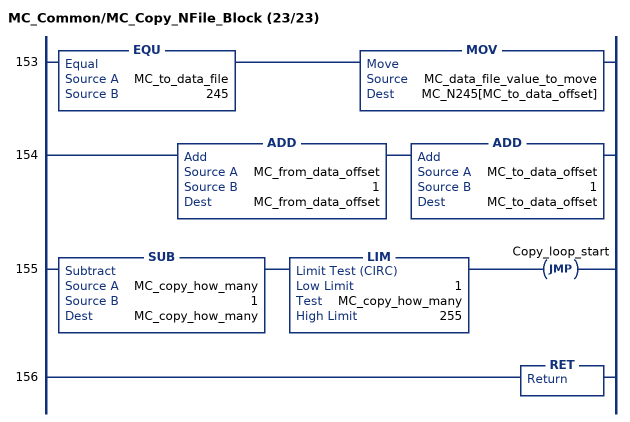
   153: EQU(MC_to_data_file,245)MOV(MC_data_file_value_to_move,MC_N245[MC_to_data_offset]);
   154: ADD(MC_from_data_offset,1,MC_from_data_offset)ADD(MC_to_data_offset,1,MC_to_data_offset);
   155: SUB(MC_copy_how_many,1,MC_copy_how_many)LIM(1,MC_copy_how_many,255)JMP(Copy_loop_start);
   156: RET();
END_ROUTINE

ROUTINE MC_DEBOUNCE_3   (* ladder *)
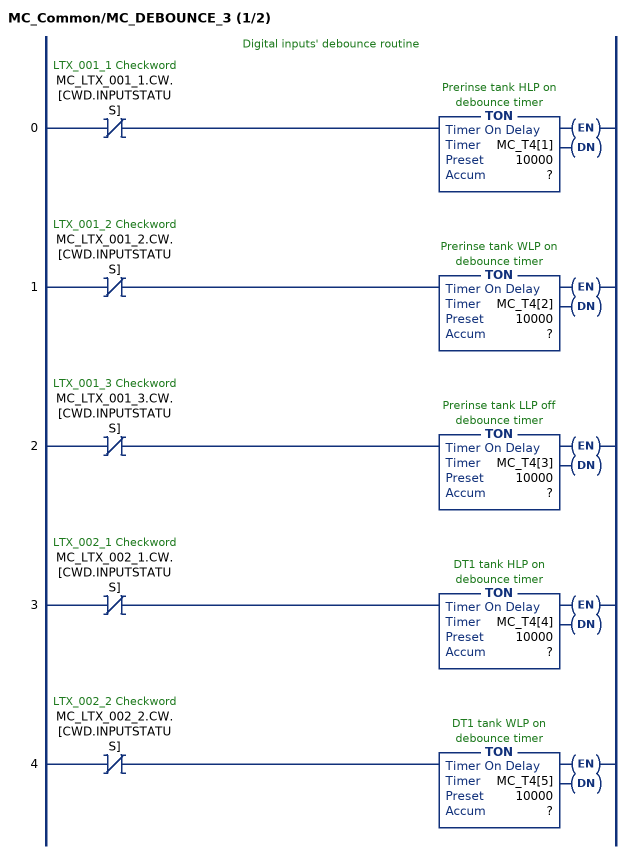
   // Digital inputs' debounce routine
   0: XIO(MC_LTX_001_1.CW.[CWD.INPUTSTATUS])TON(MC_T4[1],?,?);
   1: XIO(MC_LTX_001_2.CW.[CWD.INPUTSTATUS])TON(MC_T4[2],?,?);
   2: XIO(MC_LTX_001_3.CW.[CWD.INPUTSTATUS])TON(MC_T4[3],?,?);
   3: XIO(MC_LTX_002_1.CW.[CWD.INPUTSTATUS])TON(MC_T4[4],?,?);
   4: XIO(MC_LTX_002_2.CW.[CWD.INPUTSTATUS])TON(MC_T4[5],?,?);
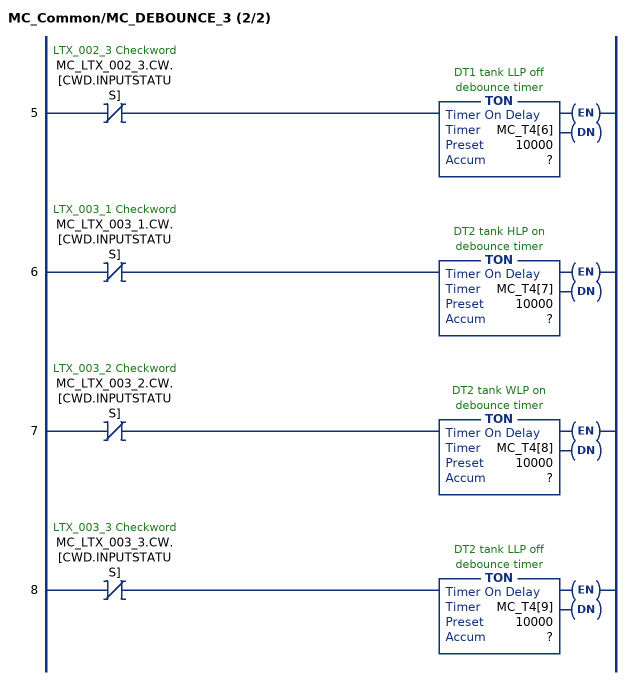
   5: XIO(MC_LTX_002_3.CW.[CWD.INPUTSTATUS])TON(MC_T4[6],?,?);
   6: XIO(MC_LTX_003_1.CW.[CWD.INPUTSTATUS])TON(MC_T4[7],?,?);
   7: XIO(MC_LTX_003_2.CW.[CWD.INPUTSTATUS])TON(MC_T4[8],?,?);
   8: XIO(MC_LTX_003_3.CW.[CWD.INPUTSTATUS])TON(MC_T4[9],?,?);
END_ROUTINE

ROUTINE MC_Digital_Inputs   (* ladder *)
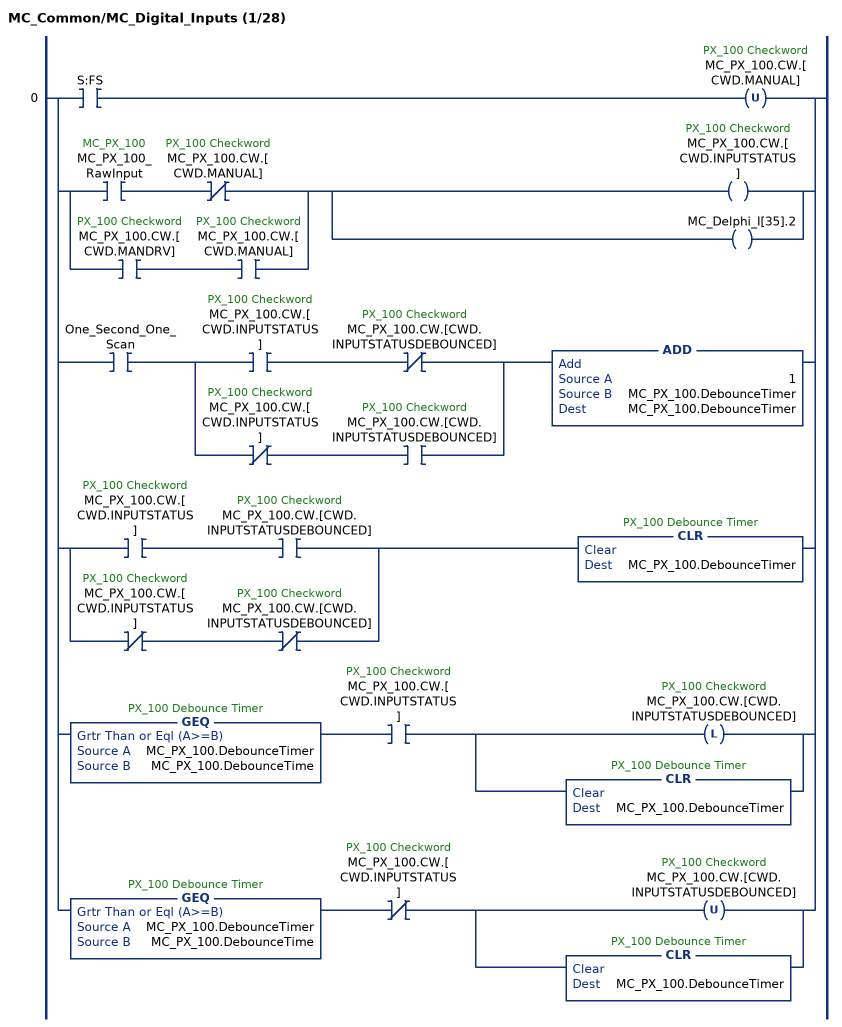
   0: [XIC(S:FS) OTU(MC_PX_100.CW.[CWD.MANUAL]) ,[XIC(MC_PX_100_RawInput) XIO(MC_PX_100.CW.[CWD.MANUAL]) ,XIC(MC_PX_100.CW.[CWD.MANDRV]) XIC(MC_PX_100.CW.[CWD.MANUAL]) ] [OTE(MC_PX_100.CW.[CWD.INPUTSTATUS]) ,OTE(MC_Delphi_I[35].2) ] ,XIC(One_Second_One_Scan) [XIC(MC_PX_100.CW.[CWD.INPUTSTATUS]) XIO(MC_PX_100.CW.[CWD.INPUTSTATUSDEBOUNCED]) ,XIO(MC_PX_100.CW.[CWD.INPUTSTATUS]) XIC(MC_PX_100.CW.[CWD.INPUTSTATUSDEBOUNCED]) ] ADD(1,MC_PX_100.DebounceTimer,MC_PX_100.DebounceTimer) ,[XIC(MC_PX_100.CW.[CWD.INPUTSTATUS]) XIC(MC_PX_100.CW.[CWD.INPUTSTATUSDEBOUNCED]) ,XIO(MC_PX_100.CW.[CWD.INPUTSTATUS]) XIO(MC_PX_100.CW.[CWD.INPUTSTATUSDEBOUNCED]) ] CLR(MC_PX_100.DebounceTimer) ,GEQ(MC_PX_100.DebounceTimer,MC_PX_100.DebounceTime) XIC(MC_PX_100.CW.[CWD.INPUTSTATUS]) [OTL(MC_PX_100.CW.[CWD.INPUTSTATUSDEBOUNCED]) ,CLR(MC_PX_100.DebounceTimer) ] ,GEQ(MC_PX_100.DebounceTimer,MC_PX_100.DebounceTime) XIO(MC_PX_100.CW.[CWD.INPUTSTATUS]) [OTU(MC_PX_100.CW.[CWD.INPUTSTATUSDEBOUNCED]) ,CLR(MC_PX_100.DebounceTimer) ] ];
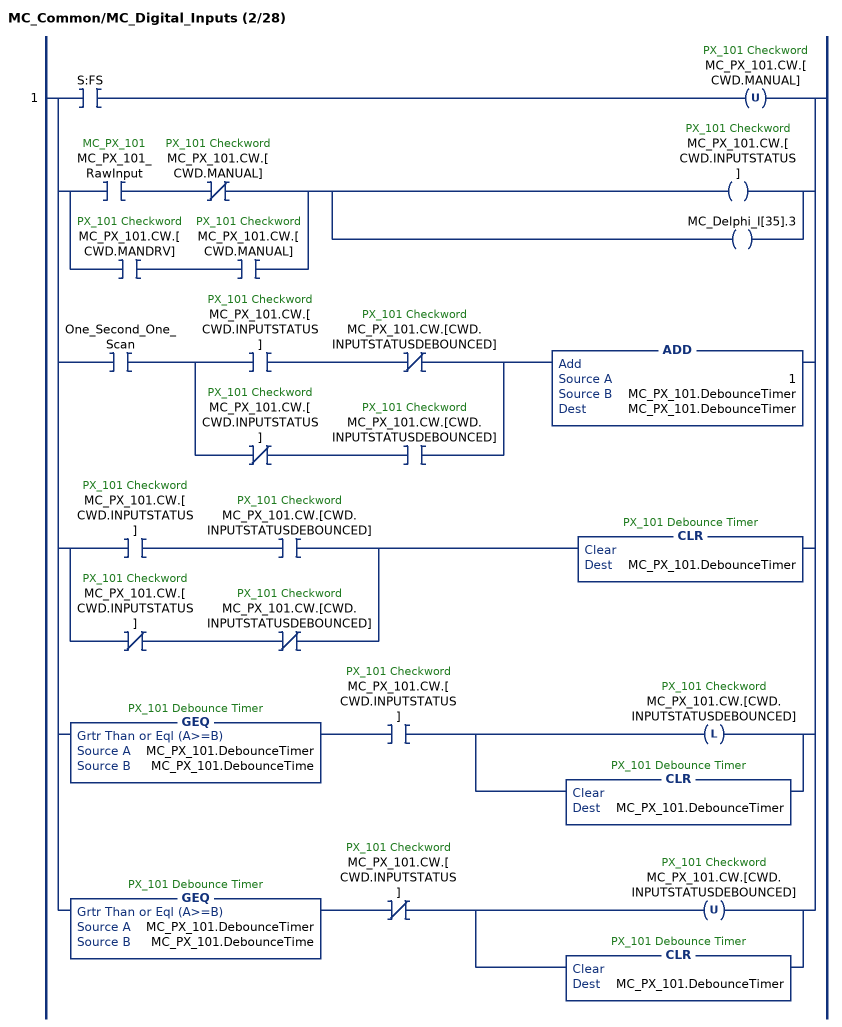
   1: [XIC(S:FS) OTU(MC_PX_101.CW.[CWD.MANUAL]) ,[XIC(MC_PX_101_RawInput) XIO(MC_PX_101.CW.[CWD.MANUAL]) ,XIC(MC_PX_101.CW.[CWD.MANDRV]) XIC(MC_PX_101.CW.[CWD.MANUAL]) ] [OTE(MC_PX_101.CW.[CWD.INPUTSTATUS]) ,OTE(MC_Delphi_I[35].3) ] ,XIC(One_Second_One_Scan) [XIC(MC_PX_101.CW.[CWD.INPUTSTATUS]) XIO(MC_PX_101.CW.[CWD.INPUTSTATUSDEBOUNCED]) ,XIO(MC_PX_101.CW.[CWD.INPUTSTATUS]) XIC(MC_PX_101.CW.[CWD.INPUTSTATUSDEBOUNCED]) ] ADD(1,MC_PX_101.DebounceTimer,MC_PX_101.DebounceTimer) ,[XIC(MC_PX_101.CW.[CWD.INPUTSTATUS]) XIC(MC_PX_101.CW.[CWD.INPUTSTATUSDEBOUNCED]) ,XIO(MC_PX_101.CW.[CWD.INPUTSTATUS]) XIO(MC_PX_101.CW.[CWD.INPUTSTATUSDEBOUNCED]) ] CLR(MC_PX_101.DebounceTimer) ,GEQ(MC_PX_101.DebounceTimer,MC_PX_101.DebounceTime) XIC(MC_PX_101.CW.[CWD.INPUTSTATUS]) [OTL(MC_PX_101.CW.[CWD.INPUTSTATUSDEBOUNCED]) ,CLR(MC_PX_101.DebounceTimer) ] ,GEQ(MC_PX_101.DebounceTimer,MC_PX_101.DebounceTime) XIO(MC_PX_101.CW.[CWD.INPUTSTATUS]) [OTU(MC_PX_101.CW.[CWD.INPUTSTATUSDEBOUNCED]) ,CLR(MC_PX_101.DebounceTimer) ] ];
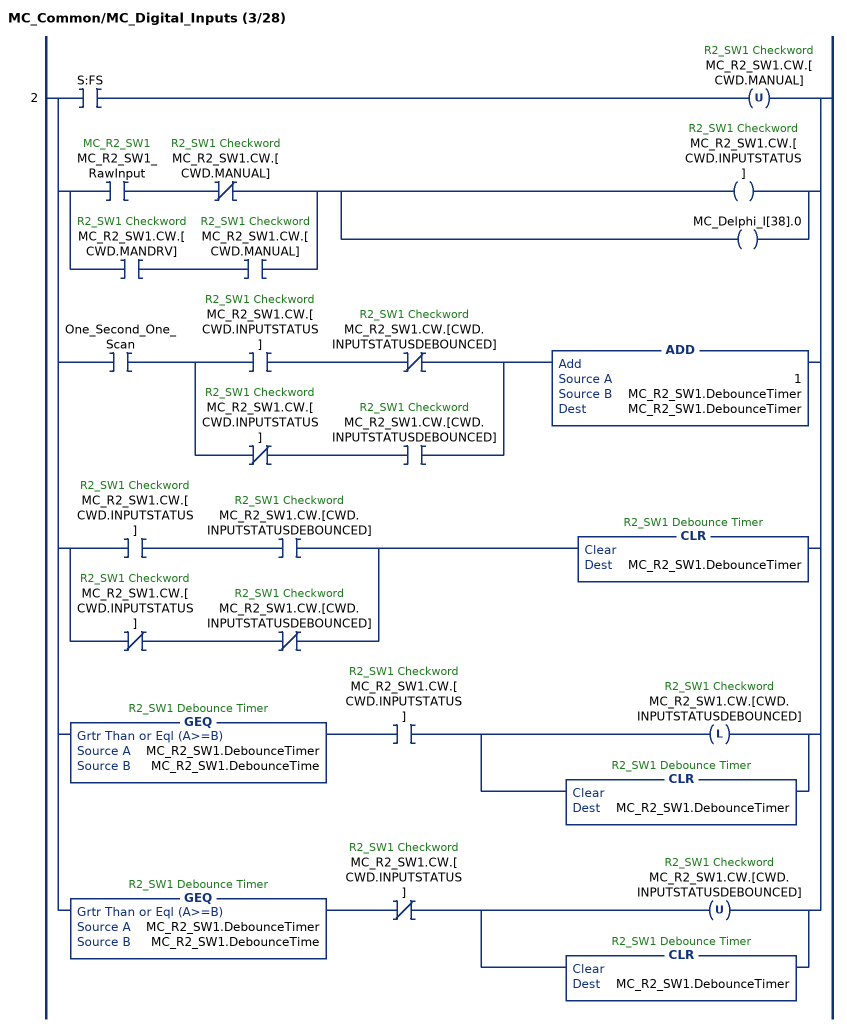
   2: [XIC(S:FS) OTU(MC_R2_SW1.CW.[CWD.MANUAL]) ,[XIC(MC_R2_SW1_RawInput) XIO(MC_R2_SW1.CW.[CWD.MANUAL]) ,XIC(MC_R2_SW1.CW.[CWD.MANDRV]) XIC(MC_R2_SW1.CW.[CWD.MANUAL]) ] [OTE(MC_R2_SW1.CW.[CWD.INPUTSTATUS]) ,OTE(MC_Delphi_I[38].0) ] ,XIC(One_Second_One_Scan) [XIC(MC_R2_SW1.CW.[CWD.INPUTSTATUS]) XIO(MC_R2_SW1.CW.[CWD.INPUTSTATUSDEBOUNCED]) ,XIO(MC_R2_SW1.CW.[CWD.INPUTSTATUS]) XIC(MC_R2_SW1.CW.[CWD.INPUTSTATUSDEBOUNCED]) ] ADD(1,MC_R2_SW1.DebounceTimer,MC_R2_SW1.DebounceTimer) ,[XIC(MC_R2_SW1.CW.[CWD.INPUTSTATUS]) XIC(MC_R2_SW1.CW.[CWD.INPUTSTATUSDEBOUNCED]) ,XIO(MC_R2_SW1.CW.[CWD.INPUTSTATUS]) XIO(MC_R2_SW1.CW.[CWD.INPUTSTATUSDEBOUNCED]) ] CLR(MC_R2_SW1.DebounceTimer) ,GEQ(MC_R2_SW1.DebounceTimer,MC_R2_SW1.DebounceTime) XIC(MC_R2_SW1.CW.[CWD.INPUTSTATUS]) [OTL(MC_R2_SW1.CW.[CWD.INPUTSTATUSDEBOUNCED]) ,CLR(MC_R2_SW1.DebounceTimer) ] ,GEQ(MC_R2_SW1.DebounceTimer,MC_R2_SW1.DebounceTime) XIO(MC_R2_SW1.CW.[CWD.INPUTSTATUS]) [OTU(MC_R2_SW1.CW.[CWD.INPUTSTATUSDEBOUNCED]) ,CLR(MC_R2_SW1.DebounceTimer) ] ];
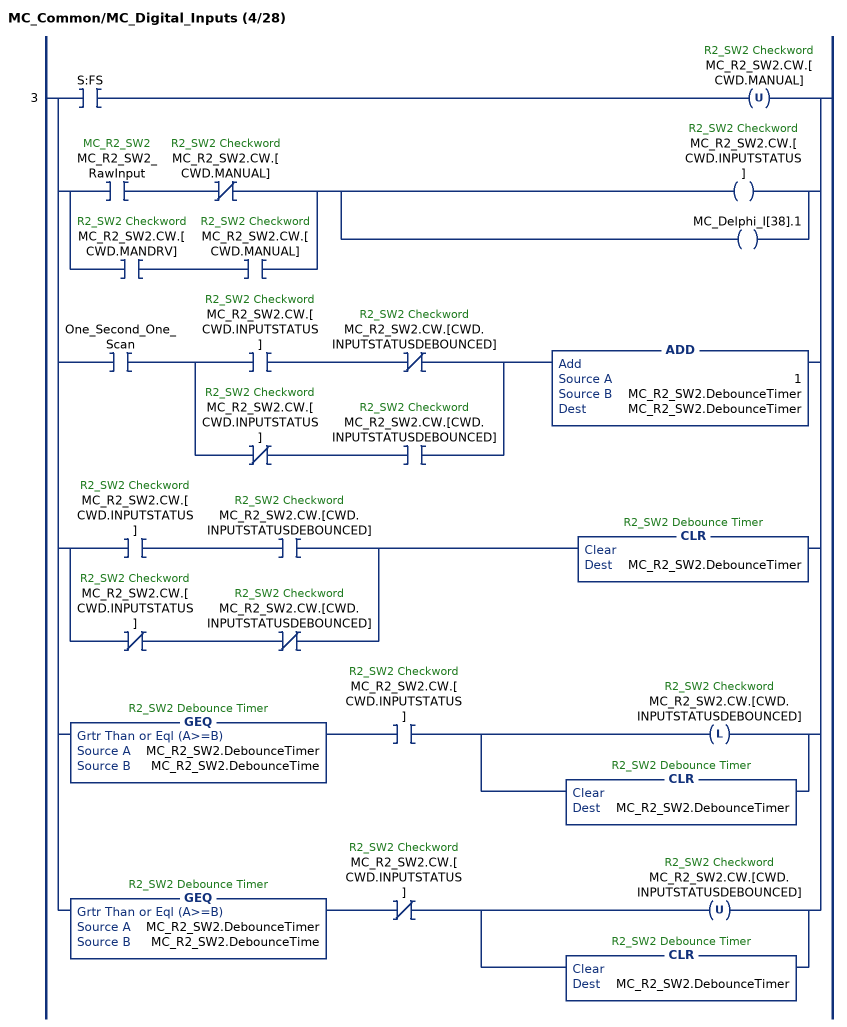
   3: [XIC(S:FS) OTU(MC_R2_SW2.CW.[CWD.MANUAL]) ,[XIC(MC_R2_SW2_RawInput) XIO(MC_R2_SW2.CW.[CWD.MANUAL]) ,XIC(MC_R2_SW2.CW.[CWD.MANDRV]) XIC(MC_R2_SW2.CW.[CWD.MANUAL]) ] [OTE(MC_R2_SW2.CW.[CWD.INPUTSTATUS]) ,OTE(MC_Delphi_I[38].1) ] ,XIC(One_Second_One_Scan) [XIC(MC_R2_SW2.CW.[CWD.INPUTSTATUS]) XIO(MC_R2_SW2.CW.[CWD.INPUTSTATUSDEBOUNCED]) ,XIO(MC_R2_SW2.CW.[CWD.INPUTSTATUS]) XIC(MC_R2_SW2.CW.[CWD.INPUTSTATUSDEBOUNCED]) ] ADD(1,MC_R2_SW2.DebounceTimer,MC_R2_SW2.DebounceTimer) ,[XIC(MC_R2_SW2.CW.[CWD.INPUTSTATUS]) XIC(MC_R2_SW2.CW.[CWD.INPUTSTATUSDEBOUNCED]) ,XIO(MC_R2_SW2.CW.[CWD.INPUTSTATUS]) XIO(MC_R2_SW2.CW.[CWD.INPUTSTATUSDEBOUNCED]) ] CLR(MC_R2_SW2.DebounceTimer) ,GEQ(MC_R2_SW2.DebounceTimer,MC_R2_SW2.DebounceTime) XIC(MC_R2_SW2.CW.[CWD.INPUTSTATUS]) [OTL(MC_R2_SW2.CW.[CWD.INPUTSTATUSDEBOUNCED]) ,CLR(MC_R2_SW2.DebounceTimer) ] ,GEQ(MC_R2_SW2.DebounceTimer,MC_R2_SW2.DebounceTime) XIO(MC_R2_SW2.CW.[CWD.INPUTSTATUS]) [OTU(MC_R2_SW2.CW.[CWD.INPUTSTATUSDEBOUNCED]) ,CLR(MC_R2_SW2.DebounceTimer) ] ];
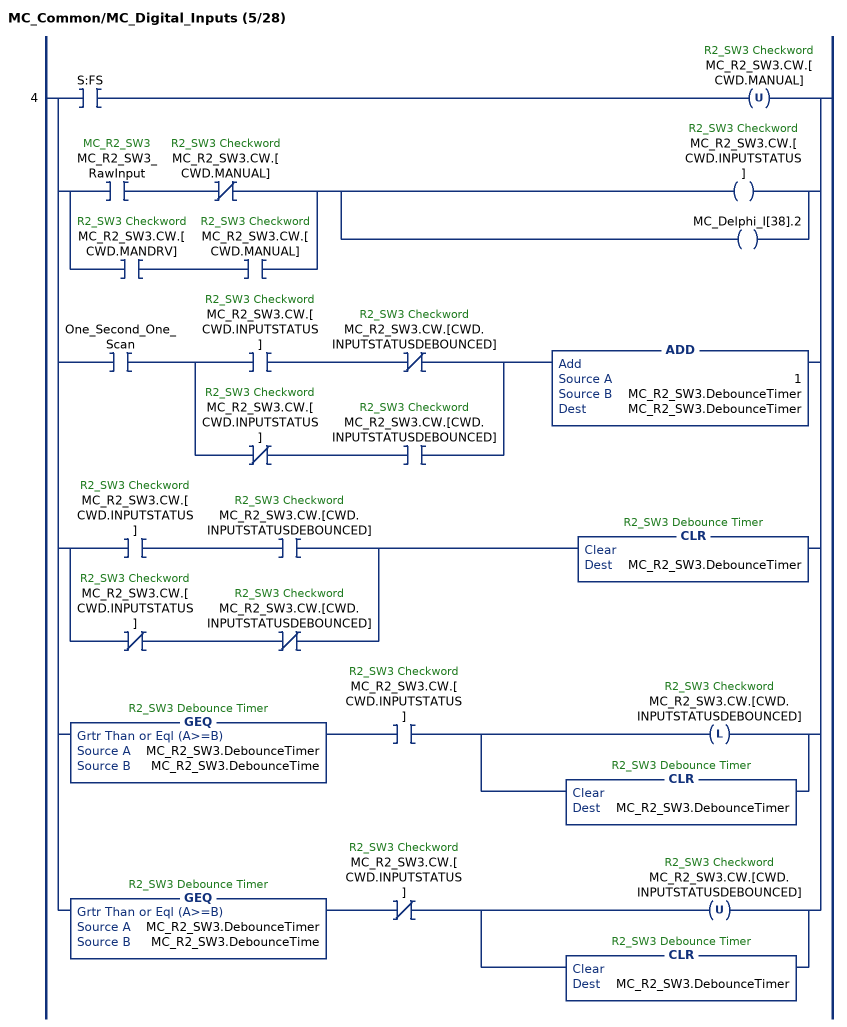
   4: [XIC(S:FS) OTU(MC_R2_SW3.CW.[CWD.MANUAL]) ,[XIC(MC_R2_SW3_RawInput) XIO(MC_R2_SW3.CW.[CWD.MANUAL]) ,XIC(MC_R2_SW3.CW.[CWD.MANDRV]) XIC(MC_R2_SW3.CW.[CWD.MANUAL]) ] [OTE(MC_R2_SW3.CW.[CWD.INPUTSTATUS]) ,OTE(MC_Delphi_I[38].2) ] ,XIC(One_Second_One_Scan) [XIC(MC_R2_SW3.CW.[CWD.INPUTSTATUS]) XIO(MC_R2_SW3.CW.[CWD.INPUTSTATUSDEBOUNCED]) ,XIO(MC_R2_SW3.CW.[CWD.INPUTSTATUS]) XIC(MC_R2_SW3.CW.[CWD.INPUTSTATUSDEBOUNCED]) ] ADD(1,MC_R2_SW3.DebounceTimer,MC_R2_SW3.DebounceTimer) ,[XIC(MC_R2_SW3.CW.[CWD.INPUTSTATUS]) XIC(MC_R2_SW3.CW.[CWD.INPUTSTATUSDEBOUNCED]) ,XIO(MC_R2_SW3.CW.[CWD.INPUTSTATUS]) XIO(MC_R2_SW3.CW.[CWD.INPUTSTATUSDEBOUNCED]) ] CLR(MC_R2_SW3.DebounceTimer) ,GEQ(MC_R2_SW3.DebounceTimer,MC_R2_SW3.DebounceTime) XIC(MC_R2_SW3.CW.[CWD.INPUTSTATUS]) [OTL(MC_R2_SW3.CW.[CWD.INPUTSTATUSDEBOUNCED]) ,CLR(MC_R2_SW3.DebounceTimer) ] ,GEQ(MC_R2_SW3.DebounceTimer,MC_R2_SW3.DebounceTime) XIO(MC_R2_SW3.CW.[CWD.INPUTSTATUS]) [OTU(MC_R2_SW3.CW.[CWD.INPUTSTATUSDEBOUNCED]) ,CLR(MC_R2_SW3.DebounceTimer) ] ];
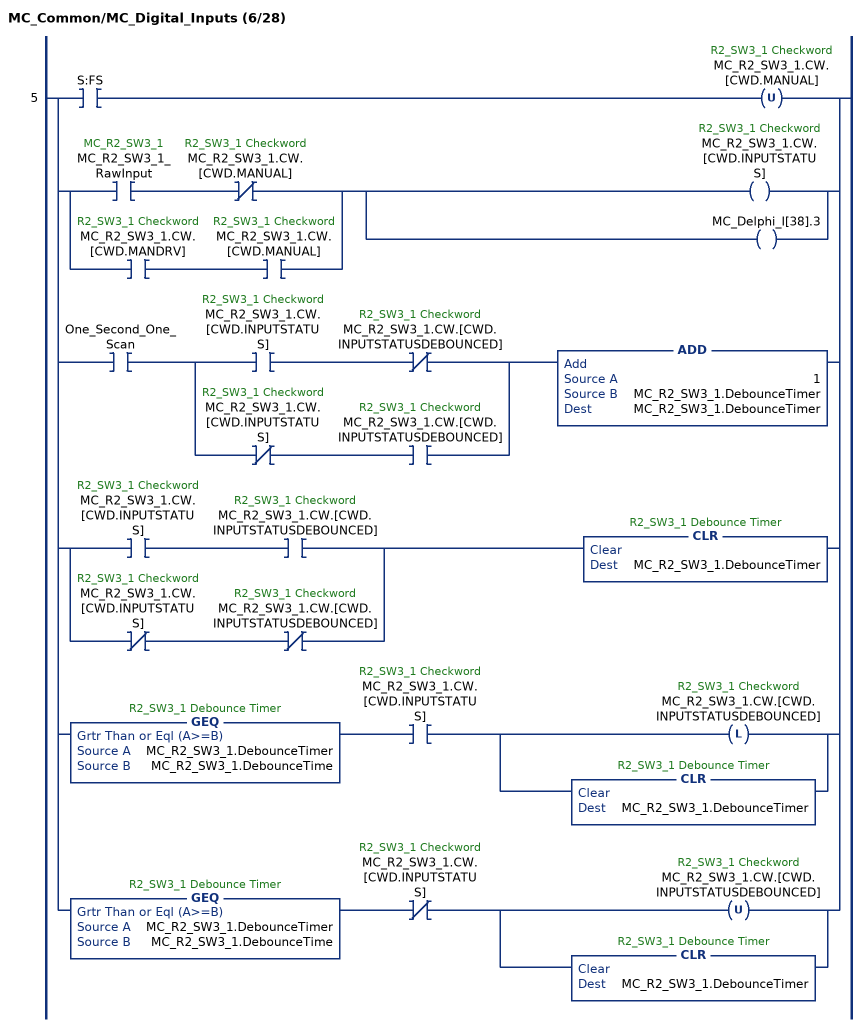
   5: [XIC(S:FS) OTU(MC_R2_SW3_1.CW.[CWD.MANUAL]) ,[XIC(MC_R2_SW3_1_RawInput) XIO(MC_R2_SW3_1.CW.[CWD.MANUAL]) ,XIC(MC_R2_SW3_1.CW.[CWD.MANDRV]) XIC(MC_R2_SW3_1.CW.[CWD.MANUAL]) ] [OTE(MC_R2_SW3_1.CW.[CWD.INPUTSTATUS]) ,OTE(MC_Delphi_I[38].3) ] ,XIC(One_Second_One_Scan) [XIC(MC_R2_SW3_1.CW.[CWD.INPUTSTATUS]) XIO(MC_R2_SW3_1.CW.[CWD.INPUTSTATUSDEBOUNCED]) ,XIO(MC_R2_SW3_1.CW.[CWD.INPUTSTATUS]) XIC(MC_R2_SW3_1.CW.[CWD.INPUTSTATUSDEBOUNCED]) ] ADD(1,MC_R2_SW3_1.DebounceTimer,MC_R2_SW3_1.DebounceTimer) ,[XIC(MC_R2_SW3_1.CW.[CWD.INPUTSTATUS]) XIC(MC_R2_SW3_1.CW.[CWD.INPUTSTATUSDEBOUNCED]) ,XIO(MC_R2_SW3_1.CW.[CWD.INPUTSTATUS]) XIO(MC_R2_SW3_1.CW.[CWD.INPUTSTATUSDEBOUNCED]) ] CLR(MC_R2_SW3_1.DebounceTimer) ,GEQ(MC_R2_SW3_1.DebounceTimer,MC_R2_SW3_1.DebounceTime) XIC(MC_R2_SW3_1.CW.[CWD.INPUTSTATUS]) [OTL(MC_R2_SW3_1.CW.[CWD.INPUTSTATUSDEBOUNCED]) ,CLR(MC_R2_SW3_1.DebounceTimer) ] ,GEQ(MC_R2_SW3_1.DebounceTimer,MC_R2_SW3_1.DebounceTime) XIO(MC_R2_SW3_1.CW.[CWD.INPUTSTATUS]) [OTU(MC_R2_SW3_1.CW.[CWD.INPUTSTATUSDEBOUNCED]) ,CLR(MC_R2_SW3_1.DebounceTimer) ] ];
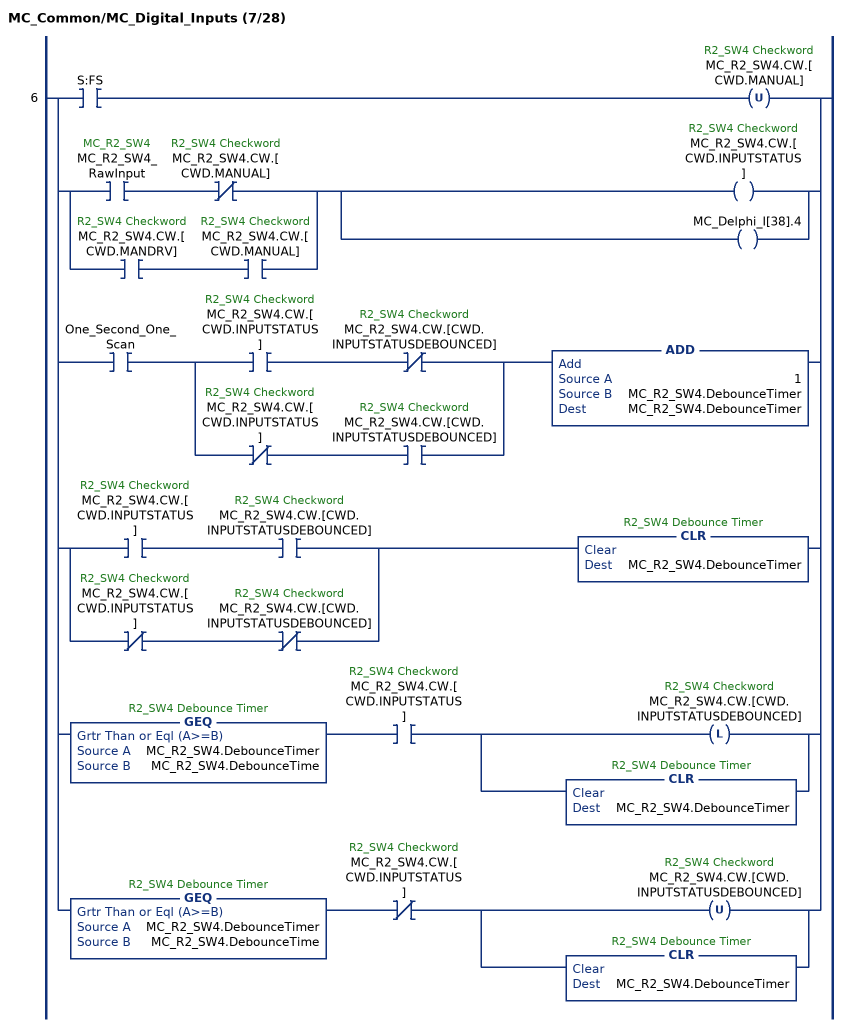
   6: [XIC(S:FS) OTU(MC_R2_SW4.CW.[CWD.MANUAL]) ,[XIC(MC_R2_SW4_RawInput) XIO(MC_R2_SW4.CW.[CWD.MANUAL]) ,XIC(MC_R2_SW4.CW.[CWD.MANDRV]) XIC(MC_R2_SW4.CW.[CWD.MANUAL]) ] [OTE(MC_R2_SW4.CW.[CWD.INPUTSTATUS]) ,OTE(MC_Delphi_I[38].4) ] ,XIC(One_Second_One_Scan) [XIC(MC_R2_SW4.CW.[CWD.INPUTSTATUS]) XIO(MC_R2_SW4.CW.[CWD.INPUTSTATUSDEBOUNCED]) ,XIO(MC_R2_SW4.CW.[CWD.INPUTSTATUS]) XIC(MC_R2_SW4.CW.[CWD.INPUTSTATUSDEBOUNCED]) ] ADD(1,MC_R2_SW4.DebounceTimer,MC_R2_SW4.DebounceTimer) ,[XIC(MC_R2_SW4.CW.[CWD.INPUTSTATUS]) XIC(MC_R2_SW4.CW.[CWD.INPUTSTATUSDEBOUNCED]) ,XIO(MC_R2_SW4.CW.[CWD.INPUTSTATUS]) XIO(MC_R2_SW4.CW.[CWD.INPUTSTATUSDEBOUNCED]) ] CLR(MC_R2_SW4.DebounceTimer) ,GEQ(MC_R2_SW4.DebounceTimer,MC_R2_SW4.DebounceTime) XIC(MC_R2_SW4.CW.[CWD.INPUTSTATUS]) [OTL(MC_R2_SW4.CW.[CWD.INPUTSTATUSDEBOUNCED]) ,CLR(MC_R2_SW4.DebounceTimer) ] ,GEQ(MC_R2_SW4.DebounceTimer,MC_R2_SW4.DebounceTime) XIO(MC_R2_SW4.CW.[CWD.INPUTSTATUS]) [OTU(MC_R2_SW4.CW.[CWD.INPUTSTATUSDEBOUNCED]) ,CLR(MC_R2_SW4.DebounceTimer) ] ];
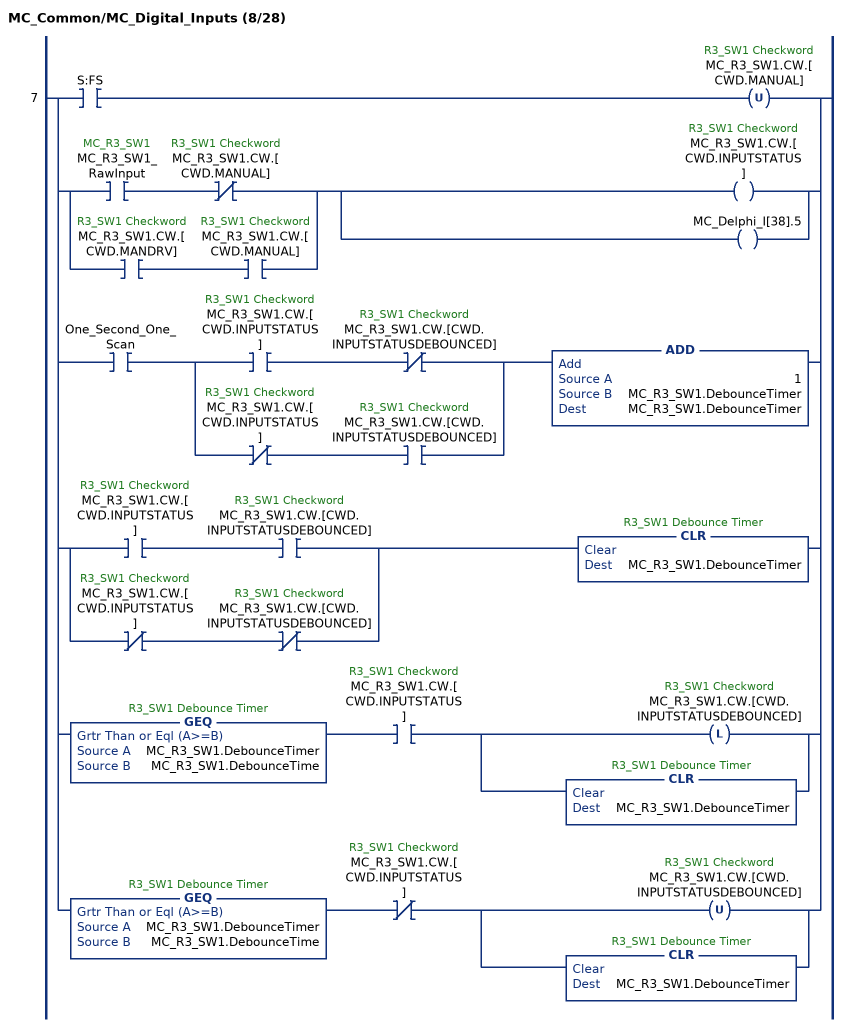
   7: [XIC(S:FS) OTU(MC_R3_SW1.CW.[CWD.MANUAL]) ,[XIC(MC_R3_SW1_RawInput) XIO(MC_R3_SW1.CW.[CWD.MANUAL]) ,XIC(MC_R3_SW1.CW.[CWD.MANDRV]) XIC(MC_R3_SW1.CW.[CWD.MANUAL]) ] [OTE(MC_R3_SW1.CW.[CWD.INPUTSTATUS]) ,OTE(MC_Delphi_I[38].5) ] ,XIC(One_Second_One_Scan) [XIC(MC_R3_SW1.CW.[CWD.INPUTSTATUS]) XIO(MC_R3_SW1.CW.[CWD.INPUTSTATUSDEBOUNCED]) ,XIO(MC_R3_SW1.CW.[CWD.INPUTSTATUS]) XIC(MC_R3_SW1.CW.[CWD.INPUTSTATUSDEBOUNCED]) ] ADD(1,MC_R3_SW1.DebounceTimer,MC_R3_SW1.DebounceTimer) ,[XIC(MC_R3_SW1.CW.[CWD.INPUTSTATUS]) XIC(MC_R3_SW1.CW.[CWD.INPUTSTATUSDEBOUNCED]) ,XIO(MC_R3_SW1.CW.[CWD.INPUTSTATUS]) XIO(MC_R3_SW1.CW.[CWD.INPUTSTATUSDEBOUNCED]) ] CLR(MC_R3_SW1.DebounceTimer) ,GEQ(MC_R3_SW1.DebounceTimer,MC_R3_SW1.DebounceTime) XIC(MC_R3_SW1.CW.[CWD.INPUTSTATUS]) [OTL(MC_R3_SW1.CW.[CWD.INPUTSTATUSDEBOUNCED]) ,CLR(MC_R3_SW1.DebounceTimer) ] ,GEQ(MC_R3_SW1.DebounceTimer,MC_R3_SW1.DebounceTime) XIO(MC_R3_SW1.CW.[CWD.INPUTSTATUS]) [OTU(MC_R3_SW1.CW.[CWD.INPUTSTATUSDEBOUNCED]) ,CLR(MC_R3_SW1.DebounceTimer) ] ];
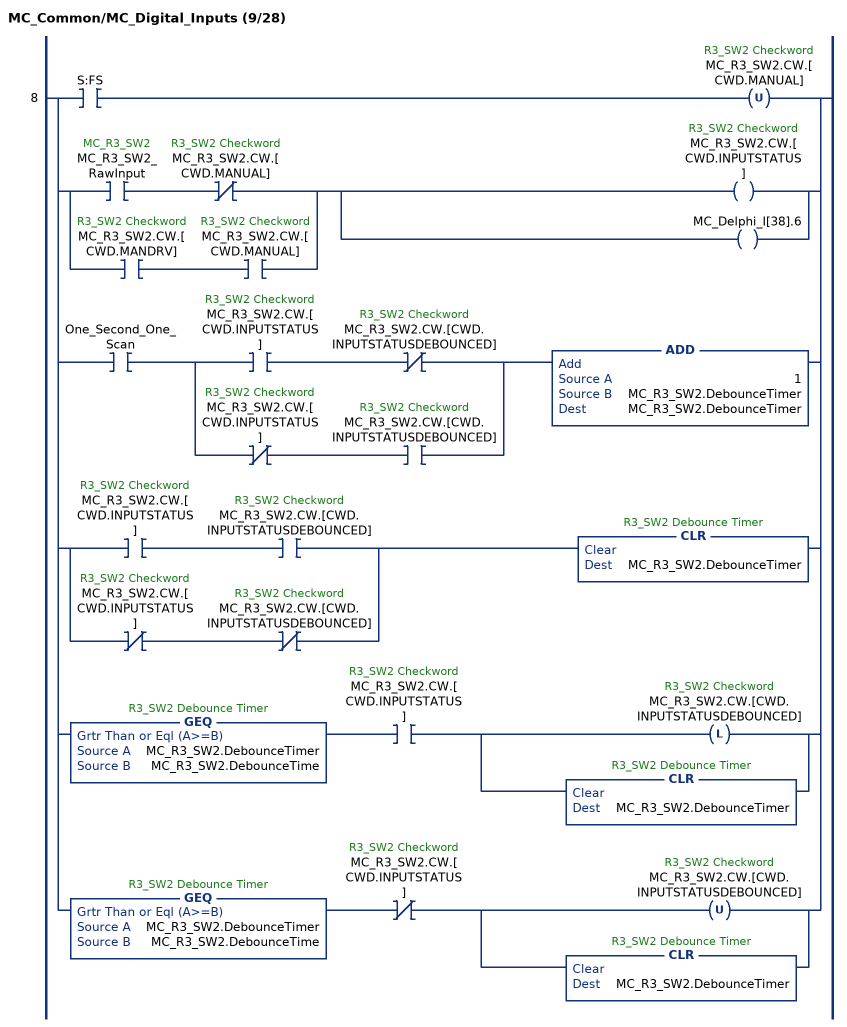
   8: [XIC(S:FS) OTU(MC_R3_SW2.CW.[CWD.MANUAL]) ,[XIC(MC_R3_SW2_RawInput) XIO(MC_R3_SW2.CW.[CWD.MANUAL]) ,XIC(MC_R3_SW2.CW.[CWD.MANDRV]) XIC(MC_R3_SW2.CW.[CWD.MANUAL]) ] [OTE(MC_R3_SW2.CW.[CWD.INPUTSTATUS]) ,OTE(MC_Delphi_I[38].6) ] ,XIC(One_Second_One_Scan) [XIC(MC_R3_SW2.CW.[CWD.INPUTSTATUS]) XIO(MC_R3_SW2.CW.[CWD.INPUTSTATUSDEBOUNCED]) ,XIO(MC_R3_SW2.CW.[CWD.INPUTSTATUS]) XIC(MC_R3_SW2.CW.[CWD.INPUTSTATUSDEBOUNCED]) ] ADD(1,MC_R3_SW2.DebounceTimer,MC_R3_SW2.DebounceTimer) ,[XIC(MC_R3_SW2.CW.[CWD.INPUTSTATUS]) XIC(MC_R3_SW2.CW.[CWD.INPUTSTATUSDEBOUNCED]) ,XIO(MC_R3_SW2.CW.[CWD.INPUTSTATUS]) XIO(MC_R3_SW2.CW.[CWD.INPUTSTATUSDEBOUNCED]) ] CLR(MC_R3_SW2.DebounceTimer) ,GEQ(MC_R3_SW2.DebounceTimer,MC_R3_SW2.DebounceTime) XIC(MC_R3_SW2.CW.[CWD.INPUTSTATUS]) [OTL(MC_R3_SW2.CW.[CWD.INPUTSTATUSDEBOUNCED]) ,CLR(MC_R3_SW2.DebounceTimer) ] ,GEQ(MC_R3_SW2.DebounceTimer,MC_R3_SW2.DebounceTime) XIO(MC_R3_SW2.CW.[CWD.INPUTSTATUS]) [OTU(MC_R3_SW2.CW.[CWD.INPUTSTATUSDEBOUNCED]) ,CLR(MC_R3_SW2.DebounceTimer) ] ];
